
screen "System screens" 1280x800, template "Template_1"
   on GenerateScreen: SetTag("Tag_ScreenNumber", 3)
   Button "Back" at 1,49 size 159x47; TextOff 'Back'
      on Release: ActivateScreen("Root screen", 0)
   Button "HmiScreenItemData" at 36,143 size 159x47; TextOff 'SIMATIC PLC system diagnos...'; PictureOff "Navigates to SIMATIC PLC system diagnostics for KTP1200 Basic+ PN 17.0.0.0"; PictureOn "Navigates to SIMATIC PLC system diagnostics for KTP1200 Basic+ PN 17.0.0.0"
      on Release: ActivateScreen("SIMATIC PLC system diagnostics", 0)
   Button "HmiScreenItemData_1" at 36,202 size 159x47; TextOff 'Project information'; PictureOff "Navigates to Project information for KTP1200 Basic+ PN 17.0.0.0"; PictureOn "Navigates to Project information for KTP1200 Basic+ PN 17.0.0.0"
      on Release: ActivateScreen("Project information", 0)
   Button "HmiScreenItemData_2" at 36,261 size 159x47; TextOff 'User administration'; PictureOff "Navigates to User administration for KTP1200 Basic+ PN 17.0.0.0"; PictureOn "Navigates to User administration for KTP1200 Basic+ PN 17.0.0.0"
      on Release: ActivateScreen("User administration", 0)
   Button "HmiScreenItemData_3" at 36,320 size 159x47; TextOff 'System information'; PictureOff "Navigates to System information for KTP1200 Basic+ PN 17.0.0.0"; PictureOn "Navigates to System information for KTP1200 Basic+ PN 17.0.0.0"
      on Release: ActivateScreen("System information", 0)
   Button "HmiScreenItemData_4" at 36,379 size 159x47; TextOff 'Different jobs'; PictureOff "Navigates to Different jobs for KTP1200 Basic+ PN 17.0.0.0"; PictureOn "Navigates to Different jobs for KTP1200 Basic+ PN 17.0.0.0"
      on Release: ActivateScreen("Different jobs", 0)

screen "SIMATIC PLC system diagnostics" 1280x800, template "Template_1"
   on GenerateScreen: SetTag("Tag_ScreenNumber", 4)
   SysDiagControl "HmiScreenItemData" at 1,97 size 1276x647
   Button "Back" at 1,49 size 159x47; TextOff 'Back'
      on Release: ActivateScreen("System screens", 0)

screen "Project information" 1280x800, template "Template_1"
   on GenerateScreen: SetTag("Tag_ScreenNumber", 5)
   TextField "HmiScreenItemData" at 35,99 size 171x28; Text 'Project name:'
   TextField "HmiScreenItemData_1" at 241,99 size 1004x28; Text 'HEAT-1-CADIZ-V5'
   TextField "HmiScreenItemData_2" at 35,129 size 171x28; Text 'Created on:'
   TextField "HmiScreenItemData_3" at 241,129 size 1004x28; Text '4/3/2025 12:55:11 PM'
   TextField "HmiScreenItemData_4" at 35,159 size 171x28; Text 'Author:'
   TextField "HmiScreenItemData_5" at 241,159 size 1004x28; Text 'User'
   TextField "HmiScreenItemData_6" at 35,189 size 171x28; Text 'Description:'
   TextField "HmiScreenItemData_7" at 241,189 size 1004x28; Text '(not configured)'
   Button "Back" at 1,49 size 159x47; TextOff 'Back'
      on Release: ActivateScreen("System screens", 0)

screen "User administration" 1280x800, template "Template_1"
   on GenerateScreen: SetTag("Tag_ScreenNumber", 6)
   UserView "HmiScreenItemData" at 1,97 size 1276x647
   Button "Back" at 1,49 size 159x47; TextOff 'Back'
      on Release: ActivateScreen("System screens", 0)

screen "System information" 1280x800, template "Template_1"
   on GenerateScreen: SetTag("Tag_ScreenNumber", 7)
   TextField "HmiScreenItemData" at 35,99 size 171x28; Text 'HMI device type:'
   TextField "HmiScreenItemData_1" at 241,99 size 1004x28; Text 'KTP1200 Basic+ PN 17.0.0.0'
   TextField "HmiScreenItemData_2" at 35,129 size 171x28; Text 'Connection:'
   TextField "HmiScreenItemData_3" at 241,129 size 1004x28; Text 'PROFINET (X1)'
   TextField "HmiScreenItemData_4" at 35,159 size 171x28; Text 'PLC:'
   TextField "HmiScreenItemData_5" at 241,159 size 1004x28; Text 'SIMATIC S7 1200'
   Button "Back" at 1,49 size 159x47; TextOff 'Back'
      on Release: ActivateScreen("System screens", 0)

screen "Different jobs" 1280x800, template "Template_1"
   on GenerateScreen: SetTag("Tag_ScreenNumber", 8)
   Button "Online" at 36,143 size 159x47; TextOff 'Online'
      on Release: function_bb44b551(0)
   Button "Offline" at 36,202 size 159x47; TextOff 'Offline'
      on Release: function_bb44b551(1)
   Button "Transfer" at 36,261 size 159x47; TextOff 'Transfer'
      on Release: function_bb44b551(2)
   Button "Toggle language" at 36,320 size 159x47; TextOff 'Toggle language'
      on Release: function_fb9197e8(-1)
   Button "Stop Runtime" at 36,379 size 159x47; TextOff 'Stop Runtime'
      on Release: StopRuntime(0)
   Button "Back" at 1,49 size 159x47; TextOff 'Back'
      on Release: ActivateScreen("System screens", 0)

screen "CUBA_FESTO_VALVULAS" 1280x800
   Switch "Switch_1" at 206,38 size 157x47; CaptionText 'Switch'; TextOff 'OFF'; TextOn 'ON'
      on SwitchOn: SetBit("HMI_CUBA_FESTO_HMI_VALVULA_52_BIESTABLE_11")
      on SwitchOff: ResetBit("HMI_CUBA_FESTO_HMI_VALVULA_52_BIESTABLE_11")
   Switch "Switch_2" at 205,165 size 157x47; CaptionText 'Switch'; TextOff 'OFF'; TextOn 'ON'
      on SwitchOn: SetBit("HMI_CUBA_FESTO_HMI_VALVULA_52_BIESTABLE_21")
      on SwitchOff: ResetBit("HMI_CUBA_FESTO_HMI_VALVULA_52_BIESTABLE_21")
   Switch "Switch_3" at 205,98 size 157x47; CaptionText 'Switch'; TextOff 'OFF'; TextOn 'ON'
      on SwitchOn: SetBit("HMI_CUBA_FESTO_HMI_VALVULA_52_BIESTABLE_12")
      on SwitchOff: ResetBit("HMI_CUBA_FESTO_HMI_VALVULA_52_BIESTABLE_12")
   Switch "Switch_4" at 205,234 size 157x47; CaptionText 'Switch'; TextOff 'OFF'; TextOn 'ON'
      on SwitchOn: SetBit("HMI_CUBA_FESTO_HMI_VALVULA_52_BIESTABLE_22")
      on SwitchOff: ResetBit("HMI_CUBA_FESTO_HMI_VALVULA_52_BIESTABLE_22")
   Switch "Switch_5" at 205,297 size 157x47; CaptionText 'Switch'; TextOff 'OFF'; TextOn 'ON'
      on SwitchOn: SetBit("HMI_CUBA_FESTO_HMI_VÁLVULA_52_MONOESTABLE_1")
      on SwitchOff: ResetBit("HMI_CUBA_FESTO_HMI_VÁLVULA_52_MONOESTABLE_1")
   Switch "Switch_6" at 205,553 size 157x47; CaptionText 'Switch'; TextOff 'OFF'; TextOn 'ON'
      on SwitchOn: SetBit("HMI_CUBA_FESTO_HMI_VÁLVULA_52_MONOESTABLE_5")
      on SwitchOff: ResetBit("HMI_CUBA_FESTO_HMI_VÁLVULA_52_MONOESTABLE_5")
   Switch "Switch_7" at 205,488 size 157x47; CaptionText 'Switch'; TextOff 'OFF'; TextOn 'ON'
      on SwitchOn: SetBit("HMI_CUBA_FESTO_HMI_VÁLVULA_52_MONOESTABLE_4")
      on SwitchOff: ResetBit("HMI_CUBA_FESTO_HMI_VÁLVULA_52_MONOESTABLE_4")
   Switch "Switch_8" at 205,361 size 157x47; CaptionText 'Switch'; TextOff 'OFF'; TextOn 'ON'
      on SwitchOn: SetBit("HMI_CUBA_FESTO_HMI_VÁLVULA_52_MONOESTABLE_2")
      on SwitchOff: ResetBit("HMI_CUBA_FESTO_HMI_VÁLVULA_52_MONOESTABLE_2")
   Switch "Switch_9" at 205,423 size 157x47; CaptionText 'Switch'; TextOff 'OFF'; TextOn 'ON'
      on SwitchOn: SetBit("HMI_CUBA_FESTO_HMI_VÁLVULA_52_MONOESTABLE_3")
      on SwitchOff: ResetBit("HMI_CUBA_FESTO_HMI_VÁLVULA_52_MONOESTABLE_3")
   TextField "Text field_1" at 28,43 size 151x32; Text 'Biestable 11'
   TextField "Text field_2" at 28,108 size 151x32; Text 'Biestable 12'
   TextField "Text field_3" at 28,177 size 151x32; Text 'Biestable 21'
   TextField "Text field_4" at 28,246 size 151x32; Text 'Biestable 22'
   TextField "Text field_5" at 9,310 size 177x32; Text 'Monoestable 1'
   TextField "Text field_6" at 9,371 size 177x32; Text 'Monoestable 2'
   TextField "Text field_7" at 14,433 size 177x32; Text 'Monoestable 3'
   TextField "Text field_8" at 19,497 size 177x32; Text 'Monoestable 4'
   TextField "Text field_9" at 17,556 size 177x32; Text 'Monoestable 5'
   Switch "Switch_10" at 612,119 size 157x47; CaptionText 'Switch'; TextOff 'OFF'; TextOn 'ON'
      on SwitchOn: SetBit("HMI_CUBA_FESTO_HMI_VÁLVULA_52_MONOESTABLE_10")
      on SwitchOff: ResetBit("HMI_CUBA_FESTO_HMI_VÁLVULA_52_MONOESTABLE_10")
   Switch "Switch_11" at 612,42 size 157x47; CaptionText 'Switch'; TextOff 'OFF'; TextOn 'ON'
      on SwitchOn: SetBit("HMI_CUBA_FESTO_HMI_VÁLVULA_52_MONOESTABLE_9")
      on SwitchOff: ResetBit("HMI_CUBA_FESTO_HMI_VÁLVULA_52_MONOESTABLE_9")
   TextField "Text field_12" at 425,49 size 177x32; Text 'Monoestable 9'
   TextField "Text field_13" at 430,118 size 192x32; Text 'Monoestable 10'
   Switch "Switch_14" at 612,408 size 157x47; CaptionText 'Switch'; TextOff 'OFF'; TextOn 'ON'
      on SwitchOn: SetBit("HMI_CUBA_FESTO_HMI_VÁLVULA_52_MONOESTABLE_14")
      on SwitchOff: ResetBit("HMI_CUBA_FESTO_HMI_VÁLVULA_52_MONOESTABLE_14")
   Switch "Switch_15" at 612,331 size 157x47; CaptionText 'Switch'; TextOff 'OFF'; TextOn 'ON'
      on SwitchOn: SetBit("HMI_CUBA_FESTO_HMI_VÁLVULA_52_MONOESTABLE_13")
      on SwitchOff: ResetBit("HMI_CUBA_FESTO_HMI_VÁLVULA_52_MONOESTABLE_13")
   Switch "Switch_16" at 612,188 size 157x47; CaptionText 'Switch'; TextOff 'OFF'; TextOn 'ON'
      on SwitchOn: SetBit("HMI_CUBA_FESTO_HMI_VÁLVULA_52_MONOESTABLE_11")
      on SwitchOff: ResetBit("HMI_CUBA_FESTO_HMI_VÁLVULA_52_MONOESTABLE_11")
   Switch "Switch_17" at 612,260 size 157x47; CaptionText 'Switch'; TextOff 'OFF'; TextOn 'ON'
      on SwitchOn: SetBit("HMI_CUBA_FESTO_HMI_VÁLVULA_52_MONOESTABLE_12")
      on SwitchOff: ResetBit("HMI_CUBA_FESTO_HMI_VÁLVULA_52_MONOESTABLE_12")
   TextField "Text field_14" at 415,200 size 192x32; Text 'Monoestable 11'
   TextField "Text field_15" at 414,269 size 192x32; Text 'Monoestable 12'
   TextField "Text field_16" at 410,336 size 192x32; Text 'Monoestable 13'
   TextField "Text field_17" at 410,408 size 192x32; Text 'Monoestable 14'
   Switch "Switch_18" at 1015,42 size 157x47; CaptionText 'Switch'; TextOff 'OFF'; TextOn 'ON'
      on SwitchOn: SetBit("HMI_CUBA_FESTO_HMI_VÁLVULA_52_MONOESTABLE_20")
      on SwitchOff: ResetBit("HMI_CUBA_FESTO_HMI_VÁLVULA_52_MONOESTABLE_20")
   TextField "Text field_21" at 824,42 size 192x32; Text 'Monoestable 20'
   Switch "Switch_22" at 1017,109 size 157x47; CaptionText 'Switch'; TextOff 'OFF'; TextOn 'ON'
      on SwitchOn: SetBit("HMI_CUBA_FESTO_HMI_VÁLVULA_52_MONOESTABLE_21")
      on SwitchOff: ResetBit("HMI_CUBA_FESTO_HMI_VÁLVULA_52_MONOESTABLE_21")
   TextField "Text field_22" at 820,121 size 192x32; Text 'Monoestable 21'
   TextField "Text field_23" at 825,190 size 192x32; Text 'Monoestable 22'
   Switch "Switch_23" at 1020,183 size 157x47; CaptionText 'Switch'; TextOff 'OFF'; TextOn 'ON'
      on SwitchOn: SetBit("HMI_CUBA_FESTO_HMI_VÁLVULA_52_MONOESTABLE_22")
      on SwitchOff: ResetBit("HMI_CUBA_FESTO_HMI_VÁLVULA_52_MONOESTABLE_22")
   TextField "Text field_24" at 409,497 size 192x32; Text 'Monoestable 15'
   Switch "Switch_24" at 619,485 size 157x47; CaptionText 'Switch'; TextOff 'OFF'; TextOn 'ON'
      on SwitchOn: SetBit("HMI_CUBA_FESTO_HMI_VÁLVULA_52_MONOESTABLE_15")
      on SwitchOff: ResetBit("HMI_CUBA_FESTO_HMI_VÁLVULA_52_MONOESTABLE_15")
   Switch "Switch_25" at 1012,337 size 157x47; CaptionText 'Switch'; TextOff 'OFF'; TextOn 'ON'
      on SwitchOn: SetBit("HMI_CUBA_FESTO_HMI_VÁLVULA_52_MONOESTABLE_24")
      on SwitchOff: ResetBit("HMI_CUBA_FESTO_HMI_VÁLVULA_52_MONOESTABLE_24")
   Switch "Switch_26" at 1017,260 size 157x47; CaptionText 'Switch'; TextOff 'OFF'; TextOn 'ON'
      on SwitchOn: SetBit("HMI_CUBA_FESTO_HMI_VÁLVULA_52_MONOESTABLE_23")
      on SwitchOff: ResetBit("HMI_CUBA_FESTO_HMI_VÁLVULA_52_MONOESTABLE_23")
   TextField "Text field_25" at 816,267 size 192x32; Text 'Monoestable 23'
   TextField "Text field_26" at 821,337 size 192x32; Text 'Monoestable 24'
   Switch "Switch_27" at 1014,404 size 157x47; CaptionText 'Switch'; TextOff 'OFF'; TextOn 'ON'
      on SwitchOn: SetBit("HMI_CUBA_FESTO_HMI_VÁLVULA_52_MONOESTABLE_25")
      on SwitchOff: ResetBit("HMI_CUBA_FESTO_HMI_VÁLVULA_52_MONOESTABLE_25")
   TextField "Text field_27" at 817,416 size 192x32; Text 'Monoestable 25'
   TextField "Text field_28" at 822,485 size 192x32; Text 'Monoestable 26'
   Switch "Switch_28" at 1027,475 size 157x47; CaptionText 'Switch'; TextOff 'OFF'; TextOn 'ON'
      on SwitchOn: SetBit("HMI_CUBA_FESTO_HMI_VÁLVULA_52_MONOESTABLE_26")
      on SwitchOff: ResetBit("HMI_CUBA_FESTO_HMI_VÁLVULA_52_MONOESTABLE_26")
   TextField "Text field_29" at 7,623 size 177x32; Text 'Monoestable 6'
   Switch "Switch_29" at 205,621 size 157x47; CaptionText 'Switch'; TextOff 'OFF'; TextOn 'ON'
      on SwitchOn: SetBit("HMI_CUBA_FESTO_HMI_VÁLVULA_52_MONOESTABLE_6")
      on SwitchOff: ResetBit("HMI_CUBA_FESTO_HMI_VÁLVULA_52_MONOESTABLE_6")
   TextField "Text field_30" at 410,550 size 192x32; Text 'Monoestable 16'
   Switch "Switch_30" at 614,547 size 157x47; CaptionText 'Switch'; TextOff 'OFF'; TextOn 'ON'
      on SwitchOn: SetBit("HMI_CUBA_FESTO_HMI_VÁLVULA_52_MONOESTABLE_16")
      on SwitchOff: ResetBit("HMI_CUBA_FESTO_HMI_VÁLVULA_52_MONOESTABLE_16")
   TextField "Text field_31" at 818,542 size 192x32; Text 'Monoestable 27'
   Switch "Switch_31" at 1016,540 size 157x47; CaptionText 'Switch'; TextOff 'OFF'; TextOn 'ON'
      on SwitchOn: SetBit("HMI_CUBA_FESTO_HMI_VÁLVULA_52_MONOESTABLE_27")
      on SwitchOff: ResetBit("HMI_CUBA_FESTO_HMI_VÁLVULA_52_MONOESTABLE_27")
   Switch "Switch_32" at 207,681 size 157x47; CaptionText 'Switch'; TextOff 'OFF'; TextOn 'ON'
      on SwitchOn: SetBit("HMI_CUBA_FESTO_HMI_VÁLVULA_52_MONOESTABLE_7")
      on SwitchOff: ResetBit("HMI_CUBA_FESTO_HMI_VÁLVULA_52_MONOESTABLE_7")
   Switch "Switch_33" at 207,753 size 157x47; CaptionText 'Switch'; TextOff 'OFF'; TextOn 'ON'
      on SwitchOn: SetBit("HMI_CUBA_FESTO_HMI_VÁLVULA_52_MONOESTABLE_8")
      on SwitchOff: ResetBit("HMI_CUBA_FESTO_HMI_VÁLVULA_52_MONOESTABLE_8")
   TextField "Text field_32" at 10,693 size 177x32; Text 'Monoestable 7'
   TextField "Text field_33" at 15,762 size 177x32; Text 'Monoestable 8'
   Switch "Switch_12" at 607,753 size 157x47; CaptionText 'Switch'; TextOff 'OFF'; TextOn 'ON'
      on SwitchOn: SetBit("HMI_CUBA_FESTO_HMI_VÁLVULA_52_MONOESTABLE_19")
      on SwitchOff: ResetBit("HMI_CUBA_FESTO_HMI_VÁLVULA_52_MONOESTABLE_19")
   Switch "Switch_13" at 607,610 size 157x47; CaptionText 'Switch'; TextOff 'OFF'; TextOn 'ON'
      on SwitchOn: SetBit("HMI_CUBA_FESTO_HMI_VÁLVULA_52_MONOESTABLE_17")
      on SwitchOff: ResetBit("HMI_CUBA_FESTO_HMI_VÁLVULA_52_MONOESTABLE_17")
   Switch "Switch_34" at 607,682 size 157x47; CaptionText 'Switch'; TextOff 'OFF'; TextOn 'ON'
      on SwitchOn: SetBit("HMI_CUBA_FESTO_HMI_VÁLVULA_52_MONOESTABLE_18")
      on SwitchOff: ResetBit("HMI_CUBA_FESTO_HMI_VÁLVULA_52_MONOESTABLE_18")
   TextField "Text field_10" at 410,622 size 192x32; Text 'Monoestable 17'
   TextField "Text field_11" at 415,691 size 192x32; Text 'Monoestable 18'
   TextField "Text field_34" at 411,760 size 192x32; Text 'Monoestable 19'
   TextField "Text field_18" at 820,610 size 192x32; Text 'Monoestable 28'
   Switch "Switch_19" at 1018,608 size 157x47; CaptionText 'Switch'; TextOff 'OFF'; TextOn 'ON'
      on SwitchOn: SetBit("HMI_CUBA_FESTO_HMI_VÁLVULA_52_MONOESTABLE_28")
      on SwitchOff: ResetBit("HMI_CUBA_FESTO_HMI_VÁLVULA_52_MONOESTABLE_28")

screen "Achim_test" 1280x800, template "Template_1"
   Switch "Switch_3" at 405,62 size 157x47; CaptionText 'Switch'; TextOff 'OFF'; TextOn 'ON'
      ProcessValue <- "hmiAchimAir"
   TextField "Text field_3" at 351,69 size 57x32; Text 'aire'
   Switch "Switch_6" at 732,66 size 157x47; CaptionText 'Switch'; TextOff 'OFF'; TextOn 'ON'
      ProcessValue <- "hmiAchimWaterInspPump"
   TextField "Text field_6" at 582,72 size 149x32; Text 'bomba agua'
   Switch "Switch_7" at 994,69 size 157x47; CaptionText 'Switch'; TextOff 'OFF'; TextOn 'ON'
      ProcessValue <- "hmiAchimInspRunning"
   TextField "Text field_7" at 936,73 size 57x32; Text 'insp'
   Button "Button_1" at 305,577 size 161x47; TextOff 'stop robot'
      on Press: SetBit("hmiAchimStopRobot")
      on Release: ResetBit("hmiAchimStopRobot")
   Button "Button_2" at 303,698 size 163x46; TextOff 'cont robot'
      on Press: SetBit("hmiAchimContRobot")
      on Release: ResetBit("hmiAchimContRobot")
   Button "Button_3" at 303,636 size 164x49; TextOff 'reset alarms'
      on Press: SetBit("hmiAchimResetAlarms")
      on Release: ResetBit("hmiAchimResetAlarms")
   GraphicIOField "PlotLight_Round_G_8" at 1023,297 size 50x50; PictureOff "PilotLight_Round_G_Off_256c"; PictureOn "PilotLight_Round_G_On_256c"
      ProcessValue <- "hmiAchimWaterInspPumpRunning"
   Switch "Switch_8" at 733,133 size 157x47; CaptionText 'Switch'; TextOff 'OFF'; TextOn 'ON'
      ProcessValue <- "hmiAchimWaterActivate"
   TextField "Text field_8" at 663,140 size 69x32; Text 'agua'
   TextField "Text field_9" at 920,367 size 97x32; Text 'agua L1'
   GraphicIOField "PlotLight_Round_G_1" at 1023,357 size 50x50; PictureOff "PilotLight_Round_G_Off_256c"; PictureOn "PilotLight_Round_G_On_256c"
      ProcessValue <- "hmiAchimWaterL1"
   TextField "Text field_10" at 922,428 size 97x32; Text 'agua L2'
   GraphicIOField "PlotLight_Round_G_2" at 1023,420 size 50x50; PictureOff "PilotLight_Round_G_Off_256c"; PictureOn "PilotLight_Round_G_On_256c"
      ProcessValue <- "hmiAchimWaterL2"
   TextField "Text field_11" at 1096,309 size 99x32; Text 'agua S1'
   GraphicIOField "PlotLight_Round_G_3" at 1199,299 size 50x50; PictureOff "PilotLight_Round_G_Off_256c"; PictureOn "PilotLight_Round_G_On_256c"
      ProcessValue <- "hmiAchimWaterS1"
   TextField "Text field_12" at 1098,370 size 99x32; Text 'agua S2'
   GraphicIOField "PlotLight_Round_G_4" at 1199,362 size 50x50; PictureOff "PilotLight_Round_G_Off_256c"; PictureOn "PilotLight_Round_G_On_256c"
      ProcessValue <- "hmiAchimWaterS2"
   TextField "Text field_13" at 1098,428 size 99x32; Text 'agua S3'
   GraphicIOField "PlotLight_Round_G_5" at 1199,420 size 50x50; PictureOff "PilotLight_Round_G_Off_256c"; PictureOn "PilotLight_Round_G_On_256c"
      ProcessValue <- "hmiAchimWaterS3"
   TextField "Text field_14" at 751,306 size 93x32; Text 'EV MPS'
   GraphicIOField "PlotLight_Round_G_6" at 852,298 size 50x50; PictureOff "PilotLight_Round_G_Off_256c"; PictureOn "PilotLight_Round_G_On_256c"
      ProcessValue <- "hmiAchimMpsEv"
   TextField "Text field_15" at 751,364 size 92x32; Text 'EV OPR'
   GraphicIOField "PlotLight_Round_G_7" at 852,356 size 50x50; PictureOff "PilotLight_Round_G_Off_256c"; PictureOn "PilotLight_Round_G_On_256c"
      ProcessValue <- "hmiAchimOprEv"
   TextField "Text field_16" at 725,424 size 125x32; Text 'antisplash'
   GraphicIOField "PlotLight_Round_G_9" at 852,416 size 50x50; PictureOff "PilotLight_Round_G_Off_256c"; PictureOn "PilotLight_Round_G_On_256c"
      ProcessValue <- "hmiAchimAntiSpash"
   TextField "Text field_17" at 567,586 size 57x32; Text 'MPS'
   GraphicIOField "PlotLight_Round_G_10" at 633,578 size 50x50; PictureOff "PilotLight_Round_G_Off_256c"; PictureOn "PilotLight_Round_G_On_256c"
      ProcessValue <- "hmiAchimMpsAlarm"
   TextField "Text field_18" at 570,644 size 57x32; Text 'OPR'
   GraphicIOField "PlotLight_Round_G_11" at 633,636 size 50x50; PictureOff "PilotLight_Round_G_Off_256c"; PictureOn "PilotLight_Round_G_On_256c"
      ProcessValue <- "hmiAchimOprAlarm"
   TextField "Text field_19" at 526,701 size 103x32; Text 'cilindros'
   GraphicIOField "PlotLight_Round_G_12" at 633,696 size 50x50; PictureOff "PilotLight_Round_G_Off_256c"; PictureOn "PilotLight_Round_G_On_256c"
      ProcessValue <- "hmiAchimPepaCylAlarm"
   TextField "Text field_20" at 794,585 size 162x32; Text 'yugo antenas'
   GraphicIOField "PlotLight_Round_G_13" at 964,578 size 50x50; PictureOff "PilotLight_Round_G_Off_256c"; PictureOn "PilotLight_Round_G_On_256c"
      ProcessValue <- "hmiAchimFrkLsAlarm"
   TextField "Text field_21" at 895,643 size 62x32; Text 'agua'
   GraphicIOField "PlotLight_Round_G_14" at 964,636 size 50x50; PictureOff "PilotLight_Round_G_Off_256c"; PictureOn "PilotLight_Round_G_On_256c"
      ProcessValue <- "hmiAchimWaterInspAlarm"
   TextField "Text field_22" at 830,698 size 129x32; Text 'agua aviso'
   GraphicIOField "PlotLight_Round_G_15" at 964,693 size 50x50; PictureOff "PilotLight_Round_G_Off_256c"; PictureOn "PilotLight_Round_G_On_256c"
      ProcessValue <- "hmiAchimWaterInspAdv"
   Button "Button_4" at 352,132 size 80x47; TextOff 'extender cilindro'
      on Press: SetBit("hmiAchimPepaCylOut")
      on Release: ResetBit("hmiAchimPepaCylOut")
   Button "Button_5" at 484,132 size 79x47; TextOff 'recoger cilindro'
      on Press: SetBit("hmiAchimPepaCylIn")
      on Release: ResetBit("hmiAchimPepaCylIn")
   TextField "Text field_4" at 933,294 size 85x60; Text 'bomba agua'
   TextField "Text field_5" at 61,298 size 108x32; Text 'acoplado'
   GraphicIOField "PlotLight_Round_G_16" at 176,294 size 50x50; PictureOff "PilotLight_Round_G_Off_256c"; PictureOn "PilotLight_Round_G_On_256c"
      ProcessValue <- "hmiAchimAirMpsCoupledE1"
   TextField "Text field_23" at 48,360 size 126x32; Text 'bloqueado'
   GraphicIOField "PlotLight_Round_G_17" at 176,352 size 50x50; PictureOff "PilotLight_Round_G_Off_256c"; PictureOn "PilotLight_Round_G_On_256c"
      ProcessValue <- "hmiAchimAirMpsLockedE2"
   TextField "Text field_24" at 8,420 size 166x32; Text 'desbloqueado'
   GraphicIOField "PlotLight_Round_G_18" at 176,412 size 50x50; PictureOff "PilotLight_Round_G_Off_256c"; PictureOn "PilotLight_Round_G_On_256c"
      ProcessValue <- "hmiAchimAirMpsUnlockedE3"
   TextField "Text field_25" at 45,479 size 129x32; Text 'presostato'
   GraphicIOField "PlotLight_Round_G_19" at 177,467 size 50x50; PictureOff "PilotLight_Round_G_Off_256c"; PictureOn "PilotLight_Round_G_On_256c"
      ProcessValue <- "hmiAchimAirMpsPressD1"
   TextField "Text field_26" at 170,255 size 57x32; Text 'MPS'
   TextField "Text field_27" at 258,252 size 162x32; Text 'antenas yugo'
   GraphicIOField "PlotLight_Round_G_20" at 381,298 size 50x50; PictureOff "PilotLight_Round_G_Off_256c"; PictureOn "PilotLight_Round_G_On_256c"
      ProcessValue <- "hmiAchimFrkLs1Nc1"
      Visibility <- "hmiAchimTool"
   GraphicIOField "PlotLight_Round_G_21" at 382,354 size 50x50; PictureOff "PilotLight_Round_G_Off_256c"; PictureOn "PilotLight_Round_G_On_256c"
      ProcessValue <- "hmiAchimFrkLs1Nc2"
      Visibility <- "hmiAchimTool"
   GraphicIOField "PlotLight_Round_G_22" at 382,411 size 50x50; PictureOff "PilotLight_Round_G_Off_256c"; PictureOn "PilotLight_Round_G_On_256c"
      ProcessValue <- "hmiAchimFrkLs2Nc1"
      Visibility <- "hmiAchimTool"
   GraphicIOField "PlotLight_Round_G_23" at 383,467 size 50x50; PictureOff "PilotLight_Round_G_Off_256c"; PictureOn "PilotLight_Round_G_On_256c"
      ProcessValue <- "hmiAchimFrkLs2Nc2"
      Visibility <- "hmiAchimTool"
   TextField "Text field_28" at 252,306 size 131x32; Text 'lado 1 NC1'
   TextField "Text field_29" at 252,360 size 131x32; Text 'lado 1 NC2'
   TextField "Text field_30" at 254,420 size 131x32; Text 'lado 2 NC1'
   TextField "Text field_31" at 254,474 size 131x32; Text 'lado 2 NC2'
   TextField "Text field_32" at 441,254 size 222x32; Text 'detectores cilindro'
   GraphicIOField "PlotLight_Round_G_24" at 598,298 size 50x50; PictureOff "PilotLight_Round_G_Off_256c"; PictureOn "PilotLight_Round_G_On_256c"
      ProcessValue <- "hmiAchimPepaCylOutProxy"
      Appearance <- "hmiAchimTool"
      Visibility <- "hmiAchimTool"
   GraphicIOField "PlotLight_Round_G_25" at 599,354 size 50x50; PictureOff "PilotLight_Round_G_Off_256c"; PictureOn "PilotLight_Round_G_On_256c"
      ProcessValue <- "hmiAchimPepaCylInProxy"
      Visibility <- "hmiAchimTool"
   TextField "Text field_33" at 475,306 size 121x32; Text 'extendido'
   TextField "Text field_34" at 487,357 size 104x32; Text 'recogido'
   TextField "Text field_35" at 927,210 size 216x37; Text 'accionamientos'
   TextField "Text field_36" at 271,209 size 149x37; Text 'detectores'
   TextField "Text field_37" at 610,531 size 113x37; Text 'alarmas'
   GraphicIOField "PlotLight_Round_G_26" at 599,464 size 50x50; PictureOff "PilotLight_Round_G_Off_256c"; PictureOn "PilotLight_Round_G_On_256c"
      ProcessValue <- "hmiAchimOprProxy"
      Visibility <- "hmiAchimTool"
   TextField "Text field_38" at 441,473 size 160x32; Text 'detector OPR'
   Switch "Switch_4" at 95,61 size 157x47; CaptionText 'Switch'; TextOff 'OFF'; TextOn 'ON'
      ProcessValue <- "hmiAchimEnable"
   TextField "Text field_39" at 1,55 size 84x60; Text 'enable HMI'
   TextField "Text field_2" at 24,125 size 58x32; Text 'tool:'
   SymbolicIOField "Symbolic I/O field_1" at 96,125 size 157x32; TextOff '0'; TextOn '1'; TextList "tool"
      ProcessValue <- "hmiAchimTool"
   TextField "Text field_1" at 22,581 size 130x32; Text '$PRO_ACT'
   GraphicIOField "PlotLight_Round_G_27" at 176,572 size 50x50; PictureOff "PilotLight_Round_G_Off_256c"; PictureOn "PilotLight_Round_G_On_256c"
      ProcessValue <- "hmiAchimPRO_ACT"
   TextField "Text field_40" at 22,639 size 147x32; Text '$STOPMESS'
   GraphicIOField "PlotLight_Round_G_28" at 176,630 size 50x50; PictureOff "PilotLight_Round_G_Off_256c"; PictureOn "PilotLight_Round_G_On_256c"
      ProcessValue <- "hmiAchimSTOPMESS"

screen "CUBA_FESTO_ENTRADAS" 1280x800
   GraphicIOField "PlotLight_Round_G" at 25,712 size 50x50; PictureOff "PilotLight_Round_G_Off_256c"; PictureOn "PilotLight_Round_G_On_256c"
      ProcessValue <- "HMI_CUBA_FESTO_HMI_SENSOR_CRDSNU_BASTIDOR_DESBLOQUEADO_2"
   GraphicIOField "PlotLight_Round_G_1" at 25,647 size 50x50; PictureOff "PilotLight_Round_G_Off_256c"; PictureOn "PilotLight_Round_G_On_256c"
      ProcessValue <- "HMI_CUBA_FESTO_HMI_SENSOR_CRDSNU_BASTIDOR_DESBLOQUEADO_1"
   GraphicIOField "PlotLight_Round_G_2" at 24,583 size 50x50; PictureOff "PilotLight_Round_G_Off_256c"; PictureOn "PilotLight_Round_G_On_256c"
      ProcessValue <- "HMI_CUBA_FESTO_HMI_SENSOR_CRDSNU_BASTIDOR_BLOQUEADO_2"
   GraphicIOField "PlotLight_Round_G_3" at 24,524 size 50x50; PictureOff "PilotLight_Round_G_Off_256c"; PictureOn "PilotLight_Round_G_On_256c"
      ProcessValue <- "HMI_CUBA_FESTO_HMI_SENSOR_CRDSNU_BASTIDOR_BLOQUEADO_1"
   GraphicIOField "PlotLight_Round_G_4" at 24,460 size 50x50; PictureOff "PilotLight_Round_G_Off_256c"; PictureOn "PilotLight_Round_G_On_256c"
      ProcessValue <- "HMI_CUBA_FESTO_HMI_Sensor_ADN_bastidor_desbloqueado_2"
   GraphicIOField "PlotLight_Round_G_5" at 24,401 size 50x50; PictureOff "PilotLight_Round_G_Off_256c"; PictureOn "PilotLight_Round_G_On_256c"
      ProcessValue <- "HMI_CUBA_FESTO_HMI_Sensor_ADN_bastidor_desbloqueado_1"
   GraphicIOField "PlotLight_Round_G_6" at 24,345 size 50x50; PictureOff "PilotLight_Round_G_Off_256c"; PictureOn "PilotLight_Round_G_On_256c"
      ProcessValue <- "HMI_CUBA_FESTO_HMI_Sensor_ADN_bastidor_bloqueado_2"
   GraphicIOField "PlotLight_Round_G_7" at 24,285 size 50x50; PictureOff "PilotLight_Round_G_Off_256c"; PictureOn "PilotLight_Round_G_On_256c"
      ProcessValue <- "HMI_CUBA_FESTO_HMI_Sensor_ADN_bastidor_bloqueado_1"
   GraphicIOField "PlotLight_Round_G_8" at 22,28 size 50x50; PictureOff "PilotLight_Round_G_Off_256c"; PictureOn "PilotLight_Round_G_On_256c"
      ProcessValue <- "HMI_CUBA_FESTO_HMI_PULSADOR_BAJAR_1"
   GraphicIOField "PlotLight_Round_G_9" at 24,225 size 50x50; PictureOff "PilotLight_Round_G_Off_256c"; PictureOn "PilotLight_Round_G_On_256c"
      ProcessValue <- "HMI_CUBA_FESTO_HMI_PULSADOR_SUBIR_2"
   GraphicIOField "PlotLight_Round_G_10" at 24,157 size 50x50; PictureOff "PilotLight_Round_G_Off_256c"; PictureOn "PilotLight_Round_G_On_256c"
      ProcessValue <- "HMI_CUBA_FESTO_HMI_PULSADOR_SUBIR_1"
   GraphicIOField "PlotLight_Round_G_11" at 24,93 size 50x50; PictureOff "PilotLight_Round_G_Off_256c"; PictureOn "PilotLight_Round_G_On_256c"
      ProcessValue <- "HMI_CUBA_FESTO_HMI_PULSADOR_BAJAR_2"
   TextField "Text field_10" at 100,34 size 186x29; Text 'Pulsador_Bajar 1'
   TextField "Text field_11" at 104,103 size 186x29; Text 'Pulsador_Bajar 2'
   TextField "Text field_12" at 108,172 size 183x29; Text 'Pulsador_Subir 1'
   TextField "Text field_13" at 112,241 size 183x29; Text 'Pulsador_Subir 2'
   TextField "Text field_14" at 104,303 size 192x29; Text 'ADN_bloqueado 1'
   TextField "Text field_15" at 106,362 size 192x29; Text 'ADN_bloqueado 2'
   TextField "Text field_16" at 106,415 size 228x29; Text 'ADN_desbloqueado 1'
   TextField "Text field_17" at 108,469 size 235x29; Text 'ADN_desbloqueado_2'
   TextField "Text field_18" at 105,537 size 391x29; Text 'CRDSNU_BASTIDOR_BLOQUEADO_1'
   TextField "Text field_19" at 103,594 size 391x29; Text 'CRDSNU_BASTIDOR_BLOQUEADO_2'
   TextField "Text field_20" at 88,656 size 433x29; Text 'CRDSNU_BASTIDOR_DESBLOQUEADO_1'
   TextField "Text field_21" at 89,722 size 433x29; Text 'CRDSNU_BASTIDOR_DESBLOQUEADO_2'
   GraphicIOField "PlotLight_Round_G_12" at 522,28 size 50x50; PictureOff "PilotLight_Round_G_Off_256c"; PictureOn "PilotLight_Round_G_On_256c"
      ProcessValue <- "HMI_CUBA_FESTO_HMI_SENSOR_DSBG_BASTIDOR_ABAJO_1"
   GraphicIOField "PlotLight_Round_G_13" at 522,287 size 50x50; PictureOff "PilotLight_Round_G_Off_256c"; PictureOn "PilotLight_Round_G_On_256c"
      ProcessValue <- "HMI_CUBA_FESTO_HMI_Sensor_plato_giro_1"
   GraphicIOField "PlotLight_Round_G_14" at 523,224 size 50x50; PictureOff "PilotLight_Round_G_Off_256c"; PictureOn "PilotLight_Round_G_On_256c"
      ProcessValue <- "HMI_CUBA_FESTO_HMI_SENSOR_DSBG_BASTIDOR_ARRIBA_2"
   GraphicIOField "PlotLight_Round_G_15" at 522,88 size 50x50; PictureOff "PilotLight_Round_G_Off_256c"; PictureOn "PilotLight_Round_G_On_256c"
      ProcessValue <- "HMI_CUBA_FESTO_HMI_SENSOR_DSBG_BASTIDOR_ABAJO_2"
   GraphicIOField "PlotLight_Round_G_16" at 522,155 size 50x50; PictureOff "PilotLight_Round_G_Off_256c"; PictureOn "PilotLight_Round_G_On_256c"
      ProcessValue <- "HMI_CUBA_FESTO_HMI_SENSOR_DSBG_BASTIDOR_ARRIBA_1"
   TextField "Text field_22" at 582,40 size 296x29; Text 'DSBG_BASTIDOR_ABAJO_1'
   TextField "Text field_23" at 575,104 size 296x29; Text 'DSBG_BASTIDOR_ABAJO_2'
   TextField "Text field_24" at 575,164 size 309x29; Text 'DSBG_BASTIDOR_ARRIBA_1'
   TextField "Text field_25" at 575,237 size 309x29; Text 'DSBG_BASTIDOR_ARRIBA_2'
   TextField "Text field_26" at 586,292 size 223x29; Text 'Sensor_plato_giro_1'
   GraphicIOField "PlotLight_Round_G_17" at 522,344 size 50x50; PictureOff "PilotLight_Round_G_Off_256c"; PictureOn "PilotLight_Round_G_On_256c"
      ProcessValue <- "HMI_CUBA_FESTO_HMI_Sensor_Plato_giro_2"
   GraphicIOField "PlotLight_Round_G_18" at 522,401 size 50x50; PictureOff "PilotLight_Round_G_Off_256c"; PictureOn "PilotLight_Round_G_On_256c"
      ProcessValue <- "HMI_CUBA_FESTO_HMI_Sensor_plato_giro_3"
   TextField "Text field_27" at 588,353 size 223x29; Text 'Sensor_plato_giro_2'
   TextField "Text field_28" at 590,414 size 223x29; Text 'Sensor_plato_giro_3'
   GraphicIOField "PlotLight_Round_G_19" at 524,463 size 50x50; PictureOff "PilotLight_Round_G_Off_256c"; PictureOn "PilotLight_Round_G_On_256c"
      ProcessValue <- "HMI_CUBA_FESTO_HMI_PULSADOR_BAJAR_4"
   GraphicIOField "PlotLight_Round_G_20" at 526,660 size 50x50; PictureOff "PilotLight_Round_G_Off_256c"; PictureOn "PilotLight_Round_G_On_256c"
      ProcessValue <- "HMI_CUBA_FESTO_HMI_PULSADOR_BAJAR_7"
   GraphicIOField "PlotLight_Round_G_21" at 526,592 size 50x50; PictureOff "PilotLight_Round_G_Off_256c"; PictureOn "PilotLight_Round_G_On_256c"
      ProcessValue <- "HMI_CUBA_FESTO_HMI_PULSADOR_BAJAR_6"
   GraphicIOField "PlotLight_Round_G_22" at 526,528 size 50x50; PictureOff "PilotLight_Round_G_Off_256c"; PictureOn "PilotLight_Round_G_On_256c"
      ProcessValue <- "HMI_CUBA_FESTO_HMI_PULSADOR_BAJAR_5"
   TextField "Text field_1" at 602,469 size 186x29; Text 'Pulsador_Bajar 4'
   TextField "Text field_2" at 606,538 size 186x29; Text 'Pulsador_Bajar 5'
   TextField "Text field_3" at 610,607 size 186x29; Text 'Pulsador_Bajar 6'
   TextField "Text field_4" at 614,676 size 186x29; Text 'Pulsador_Bajar 7'
   GraphicIOField "PlotLight_Round_G_23" at 961,27 size 50x50; PictureOff "PilotLight_Round_G_Off_256c"; PictureOn "PilotLight_Round_G_On_256c"
      ProcessValue <- "HMI_CUBA_FESTO_HMI_PULSADOR_BAJAR_8"
   GraphicIOField "PlotLight_Round_G_24" at 963,224 size 50x50; PictureOff "PilotLight_Round_G_Off_256c"; PictureOn "PilotLight_Round_G_On_256c"
      ProcessValue <- "HMI_CUBA_FESTO_HMI_PULSADOR_BAJAR_11"
   GraphicIOField "PlotLight_Round_G_25" at 963,156 size 50x50; PictureOff "PilotLight_Round_G_Off_256c"; PictureOn "PilotLight_Round_G_On_256c"
      ProcessValue <- "HMI_CUBA_FESTO_HMI_PULSADOR_BAJAR_10"
   GraphicIOField "PlotLight_Round_G_26" at 963,92 size 50x50; PictureOff "PilotLight_Round_G_Off_256c"; PictureOn "PilotLight_Round_G_On_256c"
      ProcessValue <- "HMI_CUBA_FESTO_HMI_PULSADOR_BAJAR_9"
   TextField "Text field_5" at 1039,33 size 186x29; Text 'Pulsador_Bajar 8'
   TextField "Text field_6" at 1043,102 size 186x29; Text 'Pulsador_Bajar 9'
   TextField "Text field_7" at 1047,171 size 199x29; Text 'Pulsador_Bajar 10'
   TextField "Text field_8" at 1051,240 size 196x29; Text 'Pulsador_Subir 11'
   GraphicIOField "PlotLight_Round_G_27" at 962,282 size 50x50; PictureOff "PilotLight_Round_G_Off_256c"; PictureOn "PilotLight_Round_G_On_256c"
      ProcessValue <- "HMI_CUBA_FESTO_HMI_PULSADOR_BAJAR_12"
   GraphicIOField "PlotLight_Round_G_29" at 964,411 size 50x50; PictureOff "PilotLight_Round_G_Off_256c"; PictureOn "PilotLight_Round_G_On_256c"
      ProcessValue <- "HMI_CUBA_FESTO_HMI_PULSADOR_BAJAR_14"
   GraphicIOField "PlotLight_Round_G_30" at 964,347 size 50x50; PictureOff "PilotLight_Round_G_Off_256c"; PictureOn "PilotLight_Round_G_On_256c"
      ProcessValue <- "HMI_CUBA_FESTO_HMI_PULSADOR_BAJAR_13"
   TextField "Text field_9" at 1040,288 size 199x29; Text 'Pulsador_Bajar 12'
   TextField "Text field_29" at 1044,357 size 199x29; Text 'Pulsador_Bajar 13'
   TextField "Text field_30" at 1048,426 size 199x29; Text 'Pulsador_Bajar 14'

screen "giro_auto" 1280x800, template "Template_1"
   Switch "Switch_1" at 109,144 size 64x32; CaptionText 'Switch'; TextOff 'OFF'; TextOn 'ON'
      on SwitchOn: SetBit("HMI_CUBA_FESTO_HMI_HABILITAR_AUTOMATICO")
      on SwitchOff: ResetBit("HMI_CUBA_FESTO_HMI_HABILITAR_AUTOMATICO")
   Switch "Switch_2" at 408,196 size 64x32; CaptionText 'Switch'; TextOff 'OFF'; TextOn 'ON'
   TextField "Text field_1" at 184,150 size 224x25; Text 'HABILITAR AUTOMATICO'
   Switch "Switch_3" at 407,254 size 64x32; CaptionText 'Switch'; TextOff 'OFF'; TextOn 'ON'
   Button "Button_1" at 221,196 size 146x32; TextOff 'giro positivo'
      on Press: SetBit("HMI_CUBA_FESTO_HMI_GIRO_POSITIVO_AUTO")
      on Release: ResetBit("HMI_CUBA_FESTO_HMI_GIRO_POSITIVO_AUTO")
   Button "Button_2" at 221,254 size 149x33; TextOff 'giro negativo'
      on Release: ResetBit("HMI_CUBA_FESTO_HMI_GIRO_NEGATIVO_AUTO")
      on Press: SetBit("HMI_CUBA_FESTO_HMI_GIRO_NEGATIVO_AUTO")
*)